FUNCTION_BLOCK "Flag: State Transition"   // FB4, SCL
{ S7_Optimized_Access := 'TRUE' }
VERSION : 0.1
   VAR_IN_OUT
      stns : "Station: All Stations";
   END_VAR
   VAR
      old : Struct
         stn : Array[0.."STATION_COUNT"] of Struct
            orderState : Array[0.."STATION_BUTTON_COUNT"] of Int;
         END_STRUCT;
      END_STRUCT;
   END_VAR
   VAR_TEMP
      pStn : Int;
      pBtn : Int;
      ret : Bool;
   END_VAR
BEGIN
   REGION "FOR EACH STATION"
       FOR #pStn := 0 TO "STATION_COUNT" DO

           REGION "IGNORE WIP LOAD CYCLE"
               IF NOT #stns.stn[#pStn].flags.wipSwapped THEN

                   REGION "FOR EACH BUTTON"
                       FOR #pBtn := 0 TO "STATION_BUTTON_COUNT" DO

                           REGION "RESET RETURN"
                               #ret := FALSE;
                           END_REGION

                           REGION "ON CHANGE IN STATE"
                               IF #stns.stn[#pStn].wipCmpts.orderState[#pBtn] <> #old.stn[#pStn].orderState[#pBtn] THEN

                                   REGION "SET STATE TRANSITION FLAG"
                                       #ret := true;
                                   END_REGION

                               END_IF;
                           END_REGION

                           REGION "SAVE FLAG"
                               #stns.stn[#pStn].flags.stateTransition[#pBtn] := #ret;
                           END_REGION

                       END_FOR;
                   END_REGION

               END_IF;
           END_REGION

           REGION "CHANGE DETECTION"
               #old.stn[#pStn].orderState := #stns.stn[#pStn].wipCmpts.orderState;
           END_REGION

       END_FOR;
   END_REGION
END_FUNCTION_BLOCK

FUNCTION_BLOCK "Flag"   // FB5, SCL
{ S7_Optimized_Access := 'TRUE' }
VERSION : 0.1
   VAR_INPUT
      pnLib : "Recipe: PN Text Library";
   END_VAR
   VAR_IN_OUT
      stns : "Station: All Stations";
      savedStns : "Recipe: HMI Stations Saved Wips";
   END_VAR
   VAR
      "inst New PN Code" : "Flag: New PN Code";
      "inst Flag: State Transition" : "Flag: State Transition";
      "inst Flag: Wip Deselect" : "Flag: Wip Deselect";
      "inst Flag: Wip Swapped" : "Flag: Wip Swapped";
   END_VAR
BEGIN
   REGION "NEW PART NUMBER ASSIGNED"
       #"inst New PN Code"(#stns);
   END_REGION

   REGION "PART NUMBER VALIDATION"
       "Flag: PN Good"(pnLib := #pnLib,
                       stns := #stns);
   END_REGION

   REGION "WIP SWAPPED"
       #"inst Flag: Wip Swapped"(#stns);
   END_REGION

   REGION "STATE TRANSITIONS"
       #"inst Flag: State Transition"(#stns);
   END_REGION

   REGION "WIP DESELECTION"
       #"inst Flag: Wip Deselect"(#savedStns);
   END_REGION
END_FUNCTION_BLOCK

FUNCTION_BLOCK "Flag: Wip Swapped"   // FB10, SCL
{ S7_Optimized_Access := 'TRUE' }
VERSION : 0.1
   VAR_IN_OUT
      stns : "Station: All Stations";
   END_VAR
   VAR
      old : Struct
         wipIndex : Array[0.."STATION_COUNT"] of DInt;
      END_STRUCT;
   END_VAR
   VAR_TEMP
      pStn : Int;
      ret : Bool;
   END_VAR
BEGIN
   REGION "FOR EACH STATION"
       FOR #pStn := 0 TO "STATION_COUNT" DO

           REGION "ON WIP CHANGE"
               IF #stns.stn[#pStn].wipData.index <> #old.wipIndex[#pStn] THEN

                   REGION "SET FLAG"
                       #ret := TRUE;
                   END_REGION

                   REGION "SAVE FLAG"
                       #stns.stn[#pStn].wipCmpts.flags.newPN := #ret;
                   END_REGION

               END_IF;
           END_REGION

           REGION "CHANGE DETECTION"
               #old.wipIndex[#pStn] := #stns.stn[#pStn].wipData.index;
           END_REGION

       END_FOR;
   END_REGION
END_FUNCTION_BLOCK

FUNCTION_BLOCK "Flag: Wip Deselect: Flag Pulse"   // FB17, SCL
{ S7_Optimized_Access := 'TRUE' }
VERSION : 0.1
   VAR_INPUT
      remaining : Real;
      reset : Bool;
   END_VAR
   VAR_IN_OUT
      flag : Bool;
   END_VAR
   VAR RETAIN
      hasBeenFlipped : Bool;
   END_VAR
BEGIN
   #flag := FALSE;

   IF #reset THEN
       #hasBeenFlipped := FALSE;
       RETURN;
   END_IF;

   IF #remaining >= 0.0 THEN
       #hasBeenFlipped := FALSE;
       RETURN;
   END_IF;

   IF NOT #hasBeenFlipped THEN
       IF #remaining < 0.0 THEN
           #hasBeenFlipped := TRUE;
           #flag := TRUE;
       END_IF;
   END_IF;
END_FUNCTION_BLOCK

FUNCTION_BLOCK "Flag: Wip Deselect"   // FB18, SCL
{ S7_Optimized_Access := 'TRUE' }
VERSION : 0.1
   VAR_IN_OUT
      savedStns : "Recipe: HMI Stations Saved Wips";
   END_VAR
   VAR
      "inst Flag Pulses" : Array[0.."STATION_COUNT", 0.."WIP_COUNT"] of "Flag: Wip Deselect: Flag Pulse";
   END_VAR
   VAR_TEMP
      pStn : Int;
      pWip : Int;
   END_VAR
BEGIN
   REGION "FOR EACH STATION"
       FOR #pStn := 0 TO "HMI_STATION_COUNT" DO

           REGION "FOR EACH WIP"
               FOR #pWip := 0 TO "WIP_COUNT" DO

                   REGION "FLAG PULSE"
                       #"inst Flag Pulses"[#pStn, #pWip](remaining := #savedStns.stn[#pStn].wip[#pWip].timers.wdsRemaining,
                                                         flag := #savedStns.stn[#pStn].wip[#pWip].flags.clearWipRequest);
                   END_REGION

               END_FOR;
           END_REGION

       END_FOR;
   END_REGION
END_FUNCTION_BLOCK

FUNCTION "Flag: PN Good" : Void   // FC13, SCL
{ S7_Optimized_Access := 'TRUE' }
VERSION : 0.1
   VAR_INPUT
      pnLib : "Recipe: PN Text Library";
   END_VAR
   VAR_IN_OUT
      stns : "Station: All Stations";
   END_VAR
   VAR_TEMP
      pStn : Int;
      pBtn : Int;
      pnGood : Bool;
   END_VAR
BEGIN
   REGION "FOR EACH STATION"
       FOR #pStn := 0 TO "STATION_COUNT" DO

           REGION "FOR EACH BUTTON"
               FOR #pBtn := 0 TO "STATION_BUTTON_COUNT" DO

                   REGION "ON NEW PN"
                       IF #stns.stn[#pStn].wipCmpts.flags.newPN THEN

                           REGION "VALIDATE PN"
                               #pnGood := "Validate PN"(pnCode := #stns.stn[#pStn].wipCmpts.pnCode[#pBtn],
                                                        pnLib := #pnLib);
                           END_REGION

                           REGION "SAVE TO FLAG"
                               #stns.stn[#pStn].wipCmpts.flags.pnGood[#pBtn] := #pnGood;
                           END_REGION

                       END_IF;
                   END_REGION

               END_FOR;
           END_REGION

       END_FOR;
   END_REGION
END_FUNCTION

// folder: From Excel

FUNCTION_BLOCK "From Excel"   // FB8, SCL
{ S7_Optimized_Access := 'TRUE' }
VERSION : 0.1
   VAR_INPUT
      codeLib : "From Excel: Data";
   END_VAR
   VAR_IN_OUT
      stns : "Station: All Stations";
      svdHMIStnWips : "Recipe: HMI Stations Saved Wips";
   END_VAR
   VAR
      operation_complete : Bool;
      start : Bool;
      states : "Initialize Excel Data: States";
   END_VAR
BEGIN
   REGION "STATE MACHINE"
       "Initialize Excel Data: State Machine"(start := "FirstScan" OR #start,
                                              states := #states,
                                              operation_complete := #operation_complete);
   END_REGION

   REGION "LOAD PART NUMBER CODES TO KP8 STATIONS"
       IF #states.pn_code_to_kp8_station THEN
           "From Excel: PN Code to KP8 Stations"(code_library := #codeLib,
                                                 stations := #stns,
                                                 operation_complete := #operation_complete);
       END_IF;
   END_REGION

   REGION "LOAD PART NUMBER CODES TO SAVED WIPS"
       IF #states.pn_code_to_saved_wips THEN
           "From Excel: PN Code to HMI Station Saved Wips"(code_libarary := #codeLib,
                                                           saved_wip_stations := #svdHMIStnWips,
                                                           operation_complete := #operation_complete);
       END_IF;
   END_REGION

   REGION "LOAD WIP CODES TO SAVED WIPS"
       IF #states.wip_code_to_saved_wips THEN
           "From Excel: Wip Code to HMI Station Saved WIps"(excel_code_library := #codeLib,
                                                            saved_wip_stations := #svdHMIStnWips,
                                                            operation_complete := #operation_complete);
       END_IF;
   END_REGION

   REGION "LOAD ACTIVE WIP TO HMI STATION LIST"
       IF #states.active_wip_to_hmi_station_list THEN
           "From Excel: HMI Stations Load Active WIP"(excel_code_library := #codeLib,
                                                      stations := #stns,
                                                      operation_complete := #operation_complete);
       END_IF;
   END_REGION

   REGION "LOAD ACTIVE WIP TO MASTER STATION LIST"
       IF #states.active_wip_to_master_station_list THEN
           "HMI Station: Load Active WIP into Master Station List"(operation_complete := #operation_complete);
       END_IF;
   END_REGION
END_FUNCTION_BLOCK

FUNCTION "From Excel: PN Code to KP8 Stations" : Void   // FC58, SCL
{ S7_Optimized_Access := 'TRUE' }
VERSION : 0.1
   VAR_INPUT
      code_library : "From Excel: Data";
   END_VAR
   VAR_IN_OUT
      stations : "Station: All Stations";
      operation_complete : Bool;
   END_VAR
   VAR_TEMP
      pointer_source : Int;
      pointer_destination : Int;
   END_VAR
BEGIN
   REGION "KP8 STATIONS
       FOR #pointer_source := 0 TO UDINT_TO_INT("Array.Any.Length"(#code_library.kp8Stns) - 1) DO
           #pointer_destination := #code_library.kp8Stns[#pointer_source].pStn;
           IF #pointer_destination = -1 THEN
               EXIT;
           END_IF;
           #stations.stn[#pointer_destination].wipCmpts.pnCode := #code_library.kp8Stns[#pointer_source].pnCode;
       END_FOR;
       #operation_complete := TRUE;
   END_REGION
END_FUNCTION

FUNCTION "From Excel: PN Code to HMI Station Saved Wips" : Void   // FC61, SCL
{ S7_Optimized_Access := 'TRUE' }
VERSION : 0.1
   VAR_INPUT
      code_libarary : "From Excel: Data";
   END_VAR
   VAR_IN_OUT
      saved_wip_stations : "Recipe: HMI Stations Saved Wips";
      operation_complete : Bool;
   END_VAR
   VAR_TEMP
      pointer_source_station : Int;
      pointer_destination_station : Int;
      pointer_wip : Int;
   END_VAR
BEGIN
   REGION "HMI STATIONS"
       FOR #pointer_source_station := 0 TO UDINT_TO_INT("Array.Any.Length"(#code_libarary.hmiStns) - 1) DO
           #pointer_destination_station := #code_libarary.hmiStns[#pointer_source_station].pStn;
           IF #pointer_destination_station = -1 THEN
               EXIT;
           END_IF;
           FOR #pointer_wip := 0 TO "WIP_COUNT" DO
               #saved_wip_stations.stn[#pointer_source_station].wip[#pointer_wip].pnCode :=
                   #code_libarary.hmiStns[#pointer_source_station].wip[#pointer_wip].pnCode;
           END_FOR;
       END_FOR;
       #operation_complete := TRUE;
   END_REGION
END_FUNCTION

FUNCTION "From Excel: HMI Stations Load Active WIP" : Void   // FC62, SCL
{ S7_Optimized_Access := 'TRUE' }
VERSION : 0.1
   VAR_INPUT
      excel_code_library : "From Excel: Data";
   END_VAR
   VAR_IN_OUT
      stations : "Station: All Stations";
      operation_complete : Bool;
   END_VAR
   VAR_TEMP
      pointer_source : Int;
      pointer_destination : Int;
   END_VAR
BEGIN
   REGION "HMI STATIONS"
       FOR #pointer_source := 0 TO UDINT_TO_INT("Array.Any.Length"(#excel_code_library.hmiStns) - 1) DO
           #pointer_destination := #excel_code_library.hmiStns[#pointer_source].pStn;
           IF #pointer_destination = -1 THEN
               EXIT;
           END_IF;
           #stations.stn[#pointer_destination].wipCmpts.pnCode := #excel_code_library.hmiStns[#pointer_source].wip[0].pnCode;
       END_FOR;
       #operation_complete := TRUE;
   END_REGION
END_FUNCTION

FUNCTION "From Excel: Wip Code to HMI Station Saved WIps" : Void   // FC63, SCL
{ S7_Optimized_Access := 'TRUE' }
VERSION : 0.1
   VAR_INPUT
      excel_code_library : "From Excel: Data";
   END_VAR
   VAR_IN_OUT
      saved_wip_stations : "Recipe: HMI Stations Saved Wips";
      operation_complete : Bool;
   END_VAR
   VAR_TEMP
      "pointer_source _station" : Int;
      pointer_destination_station : Int;
      pointer_wip : Int;
   END_VAR
BEGIN
   REGION "HMI STATIONS"
       FOR #"pointer_source _station" := 0 TO UDINT_TO_INT("Array.Any.Length"(#excel_code_library.hmiStns) - 1) DO
           FOR #pointer_wip := 0 TO "WIP_COUNT" DO
               #saved_wip_stations.stn[#"pointer_source _station"].wip[#pointer_wip].wip.code :=
                   #excel_code_library.hmiStns[#"pointer_source _station"].wip[#pointer_wip].wipCode;
           END_FOR;
       END_FOR;
       #operation_complete := TRUE;
   END_REGION
END_FUNCTION

FUNCTION "Initialize Excel Data: State Machine" : Void   // FC148, SCL
{ S7_Optimized_Access := 'TRUE' }
VERSION : 0.1
   VAR_INPUT
      start : Bool;
   END_VAR
   VAR_IN_OUT
      states : "Initialize Excel Data: States";
      operation_complete : Bool;
   END_VAR
   VAR_TEMP
      clear_states : "Initialize Excel Data: States";
   END_VAR
BEGIN
   REGION "LOAD PART NUMBER CODES TO KP8 STATIONS"
       IF #start AND NOT #operation_complete AND "Initialize Excel Data: All States False"(#states) THEN
           #states := #clear_states;
           #states.pn_code_to_kp8_station := TRUE;
           #operation_complete := FALSE;
       END_IF;
   END_REGION

   REGION "LOAD PART NUMBER CODES TO SAVED WIPS"
       IF #states.pn_code_to_kp8_station AND #operation_complete THEN
           #states := #clear_states;
           #states.pn_code_to_saved_wips := TRUE;
           #operation_complete := FALSE;
       END_IF;
   END_REGION

   REGION "LOAD WIP CODES TO SAVED WIPS"
       IF #states.pn_code_to_saved_wips AND #operation_complete THEN
           #states := #clear_states;
           #states.wip_code_to_saved_wips := TRUE;
           #operation_complete := FALSE;
       END_IF;
   END_REGION

   REGION "LOAD ACTIVE WIP TO HMI STATION LIST"
       IF #states.wip_code_to_saved_wips AND #operation_complete THEN
           #states := #clear_states;
           #states.active_wip_to_hmi_station_list := TRUE;
           #operation_complete := FALSE;
       END_IF;
   END_REGION

   REGION "LOAD ACTIVE WIP TO MASTER STATION LIST"
       IF #states.active_wip_to_hmi_station_list AND #operation_complete THEN
           #states := #clear_states;
           #states.active_wip_to_master_station_list := TRUE;
           #operation_complete := FALSE;
       END_IF;
   END_REGION

   REGION "COMPLETE"
       IF #states.active_wip_to_master_station_list AND #operation_complete THEN
           #states := #clear_states;
           #operation_complete := FALSE;
       END_IF;
   END_REGION
END_FUNCTION

FUNCTION "Initialize Excel Data: All States False" : Bool   // FC149, SCL
{ S7_Optimized_Access := 'TRUE' }
VERSION : 0.1
   VAR_INPUT
      states : "Initialize Excel Data: States";
   END_VAR
   VAR_TEMP
      ret : Bool;
   END_VAR
BEGIN
   IF NOT #states.active_wip_to_hmi_station_list AND
       NOT #states.pn_code_to_kp8_station AND
       NOT #states.active_wip_to_master_station_list AND
       NOT #states.pn_code_to_saved_wips AND
       NOT #states.wip_code_to_saved_wips THEN
       #ret := TRUE;
   END_IF;
   #"Initialize Excel Data: All States False" := #ret;
END_FUNCTION

// folder: Global/Physical

FUNCTION "Physical to Global" : Void   // FC1, LAD
{ S7_Optimized_Access := 'TRUE' }
VERSION : 0.1
   VAR_IN_OUT
      stations : "Station: All Stations";
   END_VAR
   VAR_TEMP
      i : Int;
      kp8In : DWord;
   END_VAR
BEGIN

REGION Network 1 (SCL): MAIN LOOP
   FOR #i := 0 TO "STATION_COUNT" DO

       CASE #i OF
           "VOLVO 16 01":
               #kp8In := "VOLVO 16 01 KP8 In";
           "VOLVO 16 02":
               #kp8In := "VOLVO 16 02 KP8 In";
           "VOLVO 16 03":
               #kp8In := "VOLVO 16 03 KP8 In";
           "VOLVO 16 04":
               #kp8In := "VOLVO 16 04 KP8 In";
           "VOLVO 16 05":
               #kp8In := "VOLVO 16 05 KP8 In";
           "VOLVO 16 06":
               #kp8In := "VOLVO 16 06 KP8 In";
           "VOLVO 16 07":
               #kp8In := "VOLVO 16 07 KP8 In";
           "VOLVO 16 08":
               #kp8In := "VOLVO 16 08 KP8 In";
           "VOLVO 16 09":
               #kp8In := "VOLVO 16 09 KP8 In";
           "VOLVO 16 10":
               #kp8In := "VOLVO 16 10 KP8 In";
           "VOLVO 16 11":
               #kp8In := "VOLVO 16 11 KP8 In";
           "CHM 01":
               #kp8In := "CHM 01 KP8 In";
           "CHM 02":
               #kp8In := "CHM 02 KP8 In";
           "CHM 03":
               #kp8In := "CHM 03 KP8 In";
           "CHM 04":
               #kp8In := "CHM 04 KP8 In";
           "CHM 05":
               #kp8In := "CHM 05 KP8 In";
           "CDO 01":
               #kp8In := "CDO 01 KP8 In";
           "CDO 02":
               #kp8In := "CDO 02 KP8 In";
           "CDO 03":
               #kp8In := "CDO 03 KP8 In";
           "BFL 01":
               #kp8In := "BFL 01 KP8 In";
           "BFL 02":
               #kp8In := "BFL 02 KP8 In";
           "BFL 03":
               #kp8In := "BFL 03 KP8 In";
           "LGS 01":
               #kp8In := "LGS 01 KP8 In";
           "LGS 02":
               #kp8In := "LGS 02 KP8 In";
           "LGS 03":
               #kp8In := "LGS 03 KP8 In";
           "CV 01":
               #kp8In := "CV 01 KP8 In";
           "CV 02":
               #kp8In := "CV 02 KP8 In";
           "CV 03":
               #kp8In := "CV 03 KP8 In";
           "CV 04":
               #kp8In := "CV 04 KP8 In";
           "PC 01":
               #kp8In := "PC 01 KP8 In"; 
           "PC 02":
               #kp8In := "PC 02 KP8 In";
       END_CASE;

       #stations.stn[#i].wipCmpts.ioData.kp8.input := #kp8In.%W1;

   END_FOR;
END_REGION
END_FUNCTION

FUNCTION "Global to Physical" : Void   // FC5, LAD
{ S7_Optimized_Access := 'TRUE' }
VERSION : 0.1
   VAR_IN_OUT
      stations : "Station: All Stations";
   END_VAR
   VAR_TEMP
      i : Int;
      j : Int;
      ET200SP : DWord;
      "KP8 In" : DWord;
      "KP8 Out" : DWord;
      Card : Int;
      stnCount : Int;
   END_VAR
BEGIN

REGION Network 1 (SCL): MAIN LOOP
   FOR #i := 0 TO "STATION_COUNT" DO

       #ET200SP := #stations.stn[#i].wipCmpts.ioData.stkLight;
       #"KP8 Out" := #stations.stn[#i].wipCmpts.ioData.kp8.tempOut;

       CASE #i OF
           "VOLVO 16 01":
               "VOLVO 16 01 IO" := #ET200SP;
               "VOLVO 16 01 KP8 Out" := #"KP8 Out";
           "VOLVO 16 02":
               "VOLVO 16 02 IO" := #ET200SP;
               "VOLVO 16 02 KP8 Out" := #"KP8 Out";
           "VOLVO 16 03":
               "VOLVO 16 03 IO" := #ET200SP;
               "VOLVO 16 03 KP8 Out" := #"KP8 Out";
           "VOLVO 16 04":
               "VOLVO 16 04 IO" := #ET200SP;
               "VOLVO 16 04 KP8 Out" := #"KP8 Out";
           "VOLVO 16 05":
               "VOLVO 16 05 IO" := #ET200SP;
               "VOLVO 16 05 KP8 Out" := #"KP8 Out";
           "VOLVO 16 06":
               "VOLVO 16 06 IO" := #ET200SP;
               "VOLVO 16 06 KP8 Out" := #"KP8 Out";
           "VOLVO 16 07":
               "VOLVO 16 07 IO" := #ET200SP;
               "VOLVO 16 07 KP8 Out" := #"KP8 Out";
           "VOLVO 16 08":
               "VOLVO 16 08 IO" := #ET200SP;
               "VOLVO 16 08 KP8 Out" := #"KP8 Out";
           "VOLVO 16 09":
               "VOLVO 16 09 IO" := #ET200SP;
               "VOLVO 16 09 KP8 Out" := #"KP8 Out";
           "VOLVO 16 10":
               "VOLVO 16 10 IO" := #ET200SP;
               "VOLVO 16 10 KP8 Out" := #"KP8 Out";
           "VOLVO 16 11":
               "VOLVO 16 11 IO" := #ET200SP;
               "VOLVO 16 11 KP8 Out" := #"KP8 Out";
           "CHM 01":
               "CHM 01 IO" := #ET200SP;
               "CHM 01 KP8 Out" := #"KP8 Out";
           "CHM 02":
               "CHM 02 IO" := #ET200SP;
               "CHM 02 KP8 Out" := #"KP8 Out";
           "CHM 03":
               "CHM 03 IO" := #ET200SP;
               "CHM 03 KP8 Out" := #"KP8 Out";
           "CHM 04":
               "CHM 04 IO" := #ET200SP;
               "CHM 04 KP8 Out" := #"KP8 Out";
           "CHM 05":
               "CHM 05 IO" := #ET200SP;
               "CHM 05 KP8 Out" := #"KP8 Out";
           "CDO 01":
               "CDO 01 IO" := #ET200SP;
               "CDO 01 KP8 Out" := #"KP8 Out";
           "CDO 02":
               "CDO 02 IO" := #ET200SP;
               "CDO 02 KP8 Out" := #"KP8 Out";
           "CDO 03":
               "CDO 03 IO" := #ET200SP;
               "CDO 03 KP8 Out" := #"KP8 Out";
           "BFL 01":
               "BFL 01 IO" := #ET200SP;
               "BFL 01 KP8 Out" := #"KP8 Out";
           "BFL 02":
               "BFL 02 IO" := #ET200SP;
               "BFL 02 KP8 Out" := #"KP8 Out";
           "BFL 03":
               "BFL 03 IO" := #ET200SP;
               "BFL 03 KP8 Out" := #"KP8 Out";
           "LGS 01":
               "LGS 01 IO" := #ET200SP;
               "LGS 01 KP8 Out" := #"KP8 Out";
           "LGS 02":
               "LGS 02 IO" := #ET200SP;
               "LGS 02 KP8 Out" := #"KP8 Out";
           "LGS 03":
               "LGS 03 IO" := #ET200SP;
               "LGS 03 KP8 Out" := #"KP8 Out";
           "CV 01":
               "CV 01 IO" := #ET200SP;
               "CV 01 KP8 Out" := #"KP8 Out";
           "CV 02":
               "CV 02 IO" := #ET200SP;
               "CV 02 KP8 Out" := #"KP8 Out";
           "CV 03":
               "CV 03 IO" := #ET200SP;
               "CV 03 KP8 Out" := #"KP8 Out";
           "CV 04":
               "CV 04 IO" := #ET200SP;
               "CV 04 KP8 Out" := #"KP8 Out";
           "PC 01":
               "PC 01 IO" := #ET200SP;
               "PC 01 KP8 Out" := #"KP8 Out";
           "PC 02":
               "PC 02 IO" := #ET200SP;
               "PC 02 KP8 Out" := #"KP8 Out";

       END_CASE;

   END_FOR;
END_REGION
END_FUNCTION

// folder: HMI: Warehouse/001 Part Call

FUNCTION_BLOCK "Part Call"   // FB16, SCL
{ S7_Optimized_Access := 'TRUE' }
VERSION : 0.1
   VAR_INPUT
      tblData : "Part Request Data";
      stns : "Station: All Stations";
      savedWips : "Recipe: HMI Stations Saved Wips";
      pnLib : "Recipe: PN Text Library";
   END_VAR
   VAR_IN_OUT
      tblHMI : "Part Call Screen";
      tableNav : "Nav Bar Data: PLC";
   END_VAR
   VAR RETAIN
      rowIndices : Array[0.."partReqTblHMIRowCnt"] of DInt;
   END_VAR
   VAR
      "inst Table Nav" : "Table Nav";
   END_VAR
   VAR_TEMP
      _tblHMI : "Part Call Screen";
      pRowHMI : DInt;
      pRowData : DInt;
   END_VAR
   // rowIndices[1] := 1;
   // rowIndices[2] := 2;
   // rowIndices[3] := 3;
   // rowIndices[4] := 4;
   // rowIndices[5] := 5;
   // rowIndices[6] := 6;
   // rowIndices[7] := 7;
   // rowIndices[8] := 8;
   // rowIndices[9] := 9;
   // rowIndices[10] := 10;
BEGIN
   REGION "TABLE NAVIGATION"
       #"inst Table Nav"(tblData := #tblData.row,
                         tblDisp := #tblHMI.row,
                         tableNav := #tableNav,
                         rowIndices := #rowIndices);
   END_REGION


   REGION "NAV BUTTON ANIMATIONS"
       "Part Call: Nav Animations"(#tableNav);
   END_REGION

   REGION "DOUBLE BUFFER IN"
       #_tblHMI := #tblHMI;
   END_REGION

   REGION "DRAW HMI TABLE"
       FOR #pRowHMI := 0 TO "partReqTblHMIRowCnt" DO

           REGION "ROW POINTER"
               #pRowData := #rowIndices[#pRowHMI];
           END_REGION

           REGION "DATA"
               "Part Call: Populate HMI Row"(address := #tblData.row[#pRowData],
                                             pnLib := #pnLib,
                                             stns := #stns,
                                             hmiRow := #_tblHMI.row[#pRowHMI]);
           END_REGION

           REGION "ANIMATIONS"
               "Part Call: Row Animations"(address := #tblData.row[#pRowData],
                                           stns := #stns,
                                           savedWips := #savedWips,
                                           rowHMI := #_tblHMI.row[#pRowHMI]);
           END_REGION

       END_FOR;
   END_REGION

   REGION "DOUBLE BUFFER OUT"
       #tblHMI := #_tblHMI;
   END_REGION
END_FUNCTION_BLOCK

FUNCTION "Part Call: Nav Animations" : Void   // FC18, SCL
{ S7_Optimized_Access := 'TRUE' }
VERSION : 0.1
   VAR_IN_OUT
      tableNav : "Nav Bar Data: PLC";
   END_VAR
   VAR_TEMP
      gray : USInt;
      green : USInt;
   END_VAR
BEGIN
   REGION "ANIMATE PART CALL NAV"

       REGION "COPY TO LOCAL"
           #gray := "GRAY_BACKGROUND";
           #green := "GREEN_LIGHT_BACKGROUND";
       END_REGION

       REGION "TOP"
           #tableNav.top.animate := "Bool.Animate"(true_color := #green,
                                                   false_color := #gray,
                                                   evaluation_signal := #tableNav.top.actuate);
       END_REGION

       REGION "PAGE UP"
           #tableNav.pageUp.animate := "Bool.Animate"(true_color := #green,
                                                      false_color := #gray,
                                                      evaluation_signal := #tableNav.pageUp.actuate);
       END_REGION

       REGION "LINE UP"
           #tableNav.lineUp.animate := "Bool.Animate"(true_color := #green,
                                                      false_color := #gray,
                                                      evaluation_signal := #tableNav.lineUp.actuate);
       END_REGION

       REGION "LINE DOWN"
           #tableNav.lineDown.animate := "Bool.Animate"(true_color := #green,
                                                        false_color := #gray,
                                                        evaluation_signal := #tableNav.lineDown.actuate);
       END_REGION

       REGION "PAGE DOWN"
           #tableNav.pageDown.animate := "Bool.Animate"(true_color := #green,
                                                        false_color := #gray,
                                                        evaluation_signal := #tableNav.pageDown.actuate);
       END_REGION

       REGION "BOTTOM"
           #tableNav.bottom.animate := "Bool.Animate"(true_color := #green,
                                                      false_color := #gray,
                                                      evaluation_signal := #tableNav.bottom.actuate);
       END_REGION

   END_REGION
END_FUNCTION

FUNCTION "Part Call: Populate HMI Row" : Void   // FC19, SCL
{ S7_Optimized_Access := 'TRUE' }
VERSION : 0.1
   VAR_INPUT
      address : DInt;
      pnLib : "Recipe: PN Text Library";
      stns : "Station: All Stations";
   END_VAR
   VAR_IN_OUT
      hmiRow : "Table Row";
   END_VAR
   VAR_TEMP
      saveAct : Bool;
      pStn : DInt;
      pWip : DInt;
      pBtn : DInt;
      blankRow : "Table Row";
   END_VAR
BEGIN
   REGION "ROW HAS DATA"
       IF #address <> -1 THEN

           REGION "GET POINTERS"
               #pStn := "Address.Get_Station"(#address);
               #pWip := "Address.Get_Wip"(#address);
               #pBtn := "Address.Get_Button"(#address);
           END_REGION

           REGION "NON WIP SPECIFIC"

           END_REGION

           REGION "GET DATA"
               #hmiRow.address := #address;
               #hmiRow.ordered := "Part Ordered"(#stns.stn[#pStn].wipCmpts.orderState[#pBtn]);
               #hmiRow.tfDropZone.value := "Strip Sign"(USINT_TO_WSTRING(#stns.stn[#pStn].id.dropZone));
               #hmiRow.tfLine.value := #stns.stn[#pStn].id.lineName;
               #hmiRow.tfPartNumber.value := "Part_Number.Code_to_WString"(pnLib := #pnLib, pnCode := #stns.stn[#pStn].wipCmpts.pnCode[#pBtn]);
               #hmiRow.tfTime.value := "Timer.Real_to_WString"(#stns.stn[#pStn].wipCmpts.timers.remaining[#pBtn]);
           END_REGION

       END_IF;
   END_REGION

   REGION "ROW HAS NO DATA"
       IF #address = -1 THEN
           #hmiRow := #blankRow;
       END_IF;
   END_REGION
END_FUNCTION

FUNCTION "Part Call: Row Animations" : Void   // FC20, SCL
{ S7_Optimized_Access := 'TRUE' }
VERSION : 0.1
   VAR_INPUT
      address : DInt;
      stns : "Station: All Stations";
      savedWips : "Recipe: HMI Stations Saved Wips";
   END_VAR
   VAR_IN_OUT
      rowHMI : "Table Row";
   END_VAR
   VAR_TEMP
      cBackground : USInt;
      cForeground : USInt;
      state : Int;
   END_VAR
BEGIN
   REGION "ROW HAS DATA"
       IF #address >= 0 THEN

           REGION "GET STATE"
               #state := "Part Call: Get State"(address := #address,
                                                stns := #stns,
                                                savedWips := #savedWips);
           END_REGION

           REGION "GET COLOR"
               "Part Call: State to Color"(state := #state,
                                           background => #cBackground,
                                           foreground => #cForeground);
           END_REGION

       END_IF;
   END_REGION

   REGION "ROW HAS NO DATA"
       IF #address <= -1 THEN
           #cForeground := "INVISIBLE";
           #cBackground := "INVISIBLE";
       END_IF;
   END_REGION


   REGION "DRAW TO HMI"
       "Part Call: Color Row"(cBackground := #cBackground,
                              cForeground := #cForeground,
                              singleLinePN := TRUE,
                              rowHMI := #rowHMI);
   END_REGION
END_FUNCTION

FUNCTION "Part Call: State to Color" : Void   // FC22, SCL
{ S7_Optimized_Access := 'TRUE' }
VERSION : 0.1
   VAR_INPUT
      state : Int;
   END_VAR
   VAR_OUTPUT
      background : USInt;
      foreground : USInt;
   END_VAR
   VAR_TEMP
      bg : USInt;
      cBlue : USInt;
      cGrayLight : USInt;
      cGrayDark : USInt;
      cGreen : USInt;
      cInvisible : USInt;
      cRedSolid : USInt;
      cRedFlash : USInt;
      cWhite : USInt;
      fg : USInt;
   END_VAR
BEGIN
   #cBlue := "BLUE_LIGHT_BACKGROUND";
   #cGreen := "GREEN_LIGHT_BACKGROUND";
   #cInvisible := "INVISIBLE";
   #cRedSolid := "RED_LIGHT_BACKGROUND";
   #cRedFlash := "RED_LIGHT_FLASHING";
   #cGrayLight := "GRAY_BACKGROUND";
   #cGrayDark := "DISABLED";
   #cWhite := "WHITE_BACKGROUND";

   CASE #state OF
       0, "idle":
           #bg := #cInvisible;
           #fg := #cInvisible;
       "requested", "acknowledged":
           #bg := #cGrayDark;
           #fg := #cGrayLight;
       "requestedCrit", "orderedCrit", "acknowledgedCrit":
           #bg := #cGrayDark;
           #fg := #cRedSolid;
       "requestedExp", "orderedExp", "acknowledgedExp":
           #bg := #cGrayDark;
           #fg := #cRedFlash;
       "ordered":
           #bg := #cGrayDark;
           #fg := #cBlue;
   END_CASE;

   #foreground := #fg;
   #background := #bg;
END_FUNCTION

FUNCTION "Part Call: Color Row" : Void   // FC31, SCL
{ S7_Optimized_Access := 'TRUE' }
VERSION : 0.1
   VAR_INPUT
      cBackground : USInt;
      cForeground : USInt;
      singleLinePN : Bool;
   END_VAR
   VAR_IN_OUT
      rowHMI : "Table Row";
   END_VAR
   VAR_TEMP
      row : "Table Row";
   END_VAR
BEGIN
   REGION "DOUBLE BUFFER IN"
       #row := #rowHMI;
   END_REGION

   REGION "INDEPENDANT ROWS"
       #row.pbSelection.animate := #cForeground;
       #row.rtBackground.animate := #cBackground;
       #row.tfDropZone.animate := #cForeground;
       #row.tfLine.animate := #cForeground;
       #row.tfTime.animate := #cForeground;
   END_REGION


   REGION "DEPENDANT ROWS"

       REGION "SINGLE LINE PART NUMBER"
           IF #singleLinePN THEN
               #row.tfPartNumber.animateDL := "INVISIBLE";
               #row.tfPartNumber.animateSL := #cForeground;
           END_IF;
       END_REGION

       REGION "DOUBLE LINE PN"
           IF NOT #singleLinePN THEN
               #row.tfPartNumber.animateDL := #cForeground;
               #row.tfPartNumber.animateSL := "INVISIBLE";
           END_IF;
       END_REGION

   END_REGION

   REGION "DOUBLE BUFFER OUT"
       #rowHMI := #row;
   END_REGION
END_FUNCTION

FUNCTION "Address in Loaded Wip" : Bool   // FC43, SCL
{ S7_Optimized_Access := 'TRUE' }
VERSION : 0.1
   VAR_INPUT
      pWip : DInt;
      stn : "Station: Single Station";
   END_VAR
   VAR_TEMP
      ret : Bool;
   END_VAR
BEGIN
   IF #pWip = #stn.wipData.index THEN
       #ret := TRUE;
   END_IF;
   #"Address in Loaded Wip" := #ret;
END_FUNCTION

FUNCTION "Part Call: Get State" : Int   // FC57, SCL
{ S7_Optimized_Access := 'TRUE' }
VERSION : 0.1
   VAR_INPUT
      address : DInt;
      stns : "Station: All Stations";
      savedWips : "Recipe: HMI Stations Saved Wips";
   END_VAR
   VAR_TEMP
      addressInWip : Bool;
      pBtn : DInt;
      pStn : DInt;
      pWip : DInt;
      ret : Int;
   END_VAR
BEGIN
   REGION "DECOMPOSE ADDRESS"
       #pBtn := "Address.Get_Button"(#address);
       #pStn := "Address.Get_Station"(#address);
       #pWip := "Address.Get_Wip"(#address);
   END_REGION

   REGION "CHECK ADDRESS AGAINST STATION'S CURRENT WIP"
       #addressInWip := "Address in Loaded Wip"(pWip := #pWip,
                                                stn := #stns.stn[#pStn]);
   END_REGION

   REGION "ADDRESS IN WIP"
       IF #addressInWip THEN
           #ret := #stns.stn[#pStn].wipCmpts.orderState[#pBtn];
       END_IF;
   END_REGION

   REGION "ADDRESS NOT IN WIP"
       IF NOT #addressInWip THEN
           #ret := #savedWips.stn[#pStn].wip[#pWip].orderState[#pBtn];
       END_IF;
   END_REGION

   REGION "RETURN"
       #"Part Call: Get State" := #ret;
   END_REGION
END_FUNCTION

// folder: HMI: Warehouse/002 Settings

FUNCTION_BLOCK "Settings Screen"   // FB19, SCL
{ S7_Optimized_Access := 'TRUE' }
VERSION : 0.1
   VAR_INPUT
      settings_meta : "Setting Meta Data";
      wip_library : "Recipe: Wip Text Library";
   END_VAR
   VAR_IN_OUT
      pn_library : "Recipe: PN Text Library";
      saved_wips : "Recipe: HMI Stations Saved Wips";
      stations : "Station: All Stations";
      settings : "Settings";
   END_VAR
   VAR
      "Assign Button" : "Assign Button";
      "Critical Time IO Field" : "Critical_IO_Field";
      "Dropzone IO Field" : "Dropzone IO Field";
      first_row : DInt;
      "Line IO Field" : "Line IO Field";
      "Part Number IO Field" : "Part Number IO Field";
      process_inputs : "Settings Screen: Processed Inputs";
      "Select Buttons Button" : "Select Buttons";
      "Select Station Button" : "Select Station PB";
      "Select WIP Button" : "Select WIP PB";
      "Table Nav_Instance" : "Table Nav";
      "Total Time IO Field" : "Total_IO_Field";
      "WIP Select Table NavBar" : "NavBar";
      inst_Selected_WIP_Table : "Selected_WIP_Table";
   END_VAR
   VAR_TEMP
      _station_rows_buffer : Array[0..2] of "Settings Station Row Data";
   END_VAR
   VAR CONSTANT
      TABLE_LENGTH : DInt := 49;
      VISIBLE_ROW_COUNT : DInt := 2;
   END_VAR
BEGIN
   REGION "SELECT STATION BUTTON"
       #"Select Station Button"(#settings.selectStation);
   END_REGION

   REGION "SELECT BUTTONS BUTTON"
       #"Select Buttons Button"(settings_meta := #settings_meta,
                                stations := #stations,
                                interface := #settings.selectButton);
   END_REGION

   REGION "SELECT WIP BUTTON"
       #"Select WIP Button"(settings_meta := #settings_meta,
                            stations := #stations,
                            interface := #settings.selectWip);
   END_REGION

   REGION "LINE IO FIELD"
       #"Line IO Field"(settings_meta := #settings_meta,
                        stations := #stations,
                        interface := #settings.line,
                        get_line := #process_inputs.line_name);
   END_REGION

   REGION "DROPZONE IO FIELD"
       #"Dropzone IO Field"(settings_meta := #settings_meta,
                            stations := #stations,
                            interface := #settings.dropzone,
                            get_dropzone := #process_inputs.dropzone);
   END_REGION

   REGION "TOTAL TIME IO FIELD"
       #"Total Time IO Field"(settings_meta := #settings_meta,
                              stations := #stations,
                              interface := #settings.total,
                              state_changes := #process_inputs.total);
   END_REGION

   REGION "CRITICAL TIME IO FIELD"
       #"Critical Time IO Field"(settings_meta := #settings_meta,
                                 stations := #stations,
                                 interface := #settings.critical,
                                 state_changes := #process_inputs.critical);
   END_REGION

   REGION "PART NUMBER ENTRY FIELD"
       #"Part Number IO Field"(settings_meta := #settings_meta,
                               stations := #stations,
                               interface := #settings.partNumber,
                               get_part_number := #process_inputs.part_number_single);

   END_REGION

   REGION "ASSIGN BUTTON"
       #"Assign Button"(critical_time := #settings.critical,
                        drop_zone := #settings.dropzone,
                        line := #settings.line,
                        part_number := #settings.partNumber,
                        settings_meta := #settings_meta,
                        total_time := #settings.total,
                        pn_library := #pn_library,
                        saved_wips := #saved_wips,
                        stations := #stations,
                        interface := #settings.assign,
                        state_changes := #process_inputs.assign);
   END_REGION

   REGION "SELECTED WIP TABLE"
       #_station_rows_buffer := #settings.stationRows;
       #inst_Selected_WIP_Table(saved_wips := #saved_wips,
                                settings_meta := #settings_meta,
                                stations := #stations,
                                wip_library := #wip_library,
                                pn_library := #pn_library,
                                navigation_bar := #settings.stnTableNavBar.plc,
                                stationRows := #_station_rows_buffer);
       #settings.stationRows := #_station_rows_buffer;
   END_REGION

   REGION "WIP SELECT TABLE NAVBAR"
       #"WIP Select Table NavBar"(hide := #settings_meta.selected_stations.count < 4,
                                  TABLE_LENGTH := #TABLE_LENGTH,
                                  VISIBLE_ROW_COUNT := #VISIBLE_ROW_COUNT,
                                  interface := #settings.stnTableNavBar,
                                  first_row := #first_row);
   END_REGION
END_FUNCTION_BLOCK

FUNCTION "Settings Screen: Load Selected: Non-HMI Station" : Void   // FC150, SCL
{ S7_Optimized_Access := 'TRUE' }
VERSION : 0.1
   VAR_INPUT
      stations : "Station: All Stations";
      selected_stations : "Selected Stations";
      wip_library : "Recipe: Wip Text Library";
      part_number_library : "Recipe: PN Text Library";
   END_VAR
   VAR_IN_OUT
      selected_station_table : Array[0..2] of "Settings Station Row Data";
   END_VAR
   VAR_TEMP
      station_index : Int;
      table_row_index : Int;
   END_VAR
BEGIN
   FOR #station_index := 0 TO "STATION_COUNT" DO
       IF #selected_stations.stns[#station_index] THEN
           "Settings Screen: Load Selected WIP"(station := #stations.stn[#station_index],
                                                wip_library := #wip_library,
                                                part_number_library := #part_number_library,
                                                table_row := #selected_station_table[#table_row_index]);
           #table_row_index += 1;
           IF #table_row_index > 2 THEN
               EXIT;
           END_IF;
       END_IF;
   END_FOR;
END_FUNCTION

FUNCTION "Settings Screen: Load Selected WIP" : Void   // FC151, SCL
{ S7_Optimized_Access := 'TRUE' }
VERSION : 0.1
   VAR_INPUT
      station : "Station: Single Station";
      wip_library : "Recipe: Wip Text Library";
      part_number_library : "Recipe: PN Text Library";
   END_VAR
   VAR_IN_OUT
      table_row : "Settings Station Row Data";
   END_VAR
   VAR_TEMP
      _table_row : "Settings Station Row Data";
      button_index : Int;
   END_VAR
BEGIN
   REGION "NOTES"
       (*
       Simple data map from station presented at input to hmi data structure.
       Decision about which data to map is done in parent.
       last edit: 2021-10-06
       *)
   END_REGION

   REGION "BUFFER IN"
       #_table_row := #table_row;
   END_REGION

   REGION "MAP"
       #_table_row.line.data := #station.id.lineName;
       #_table_row.dropzone.data := "Strip Sign"(USINT_TO_WSTRING(#station.id.dropZone));
       #_table_row.wip.data := "WIP.Code_to_WString"(wipTxtLib := #wip_library,
                                                           code := #station.wipData.code);
       FOR #button_index := 0 TO "STATION_BUTTON_COUNT" DO
           "Settings Screen: Load Selected WIP: Load Button"(wip_components:=#station.wipCmpts,
                                                                 wip_library := #wip_library,
                                                                 button_index := #button_index,
                                                                 part_number_liberary := #part_number_library,
                                                                 button_row := #_table_row.btnRows[#button_index]);
       END_FOR;
   END_REGION

   REGION "BUFFER OUT"
       #table_row := #_table_row;
   END_REGION
END_FUNCTION

FUNCTION "Settings Screen: Selected Station Table Row Color" : Void   // FC152, SCL
{ S7_Optimized_Access := 'TRUE' }
VERSION : 0.1
BEGIN
END_FUNCTION

FUNCTION "Settings Screen: Load Selected WIP: Load Button" : Void   // FC155, SCL
{ S7_Optimized_Access := 'TRUE' }
VERSION : 0.1
   VAR_INPUT
      button_index : Int;
      part_number_liberary : "Recipe: PN Text Library";
      wip_components : "Station: Wip: Wip Module";
      wip_library : "Recipe: Wip Text Library";
   END_VAR
   VAR_IN_OUT
      button_row : "Settings Station Row Button Row Data";
   END_VAR
   VAR_TEMP
      _button_row : "Settings Station Row Button Row Data";
      part_number_wstring : WString;
      part_number_code : DInt;
   END_VAR
   VAR CONSTANT
      no_code : WString;
   END_VAR
BEGIN
   REGION "NOTES"
       (*
       Simple data map from station presented at input to hmi data structure.
       Decision about which data to map is done in parent.
       last edit: 2021-10-06
       *)
   END_REGION

   REGION "BUFFER IN"    
       #_button_row := #button_row;
   END_REGION

   REGION "BUTTON LABEL"
       // CURRENTLY A STATIC LABEL
   END_REGION

   REGION "ALOTTED TIME"
       #_button_row.total.data := "Timer.Real_to_WString"(#wip_components.timers.ptAllotted[#button_index]);
   END_REGION

   REGION "CRITICAL TIME"
       #_button_row.critical.data := "Timer.Real_to_WString"(#wip_components.timers.ptCritical[#button_index]);
   END_REGION

   REGION "PART NUMBER"

       REGION "PROCESS PART NUMBER"
           #part_number_code := #wip_components.pnCode[#button_index];
           #part_number_wstring := "Part_Number.Code_to_WString"(pnLib := #part_number_liberary,
                                                         pnCode := #part_number_code);
       END_REGION

       REGION "SINGLE LINE PART NUMBER"
           IF "Part_Number.Is_Single"(#part_number_code) THEN
               #_button_row.singlePN.data := #part_number_wstring;
               #_button_row.doublePN.data := #no_code;
           END_IF;
       END_REGION

       REGION "DOUBLE LINE PART NUMBER"
           IF "Part_Number.Is_Double"(#part_number_code) THEN
               #_button_row.singlePN.data := #no_code;
               #_button_row.doublePN.data := #part_number_wstring;
           END_IF;
       END_REGION

   END_REGION

   REGION "BUFFER OUT"
       #button_row := #_button_row;
   END_REGION
END_FUNCTION

FUNCTION "Settings Screen: Load Selected: HMI Station" : Void   // FC176, SCL
{ S7_Optimized_Access := 'TRUE' }
VERSION : 0.1
   VAR_INPUT
      stations : "Station: All Stations";
      selected_wips : "Selected Wips";
      wip_library : "Recipe: Wip Text Library";
      part_number_library : "Recipe: PN Text Library";
   END_VAR
   VAR_IN_OUT
      selected_station_table : Array[0..2] of "Settings Station Row Data";
   END_VAR
   VAR_TEMP
      station_index : Int;
      table_row_index : Int;
   END_VAR
BEGIN
   FOR #station_index := 0 TO #selected_wips.count DO
       "Settings Screen: Load Selected WIP"(station := #stations.stn[#station_index],
                                            wip_library := #wip_library,
                                            part_number_library := #part_number_library,
                                            table_row := #selected_station_table[#table_row_index]);END_FOR;
END_FUNCTION

// folder: HMI: Warehouse/002 Settings/Assign Button

FUNCTION_BLOCK "Assign Button"   // FB55, SCL
{ S7_Optimized_Access := 'TRUE' }
VERSION : 0.1
   VAR_INPUT
      critical_time : "IO Field Data: Label with Data";
      drop_zone : "IO Field Data: Label with Data";
      line : "IO Field Data: Label with Data";
      part_number : "IO Field Data: Label with Data";
      settings_meta : "Setting Meta Data";
      total_time : "IO Field Data: Label with Data";
   END_VAR
   VAR_IN_OUT
      interface : "Push Button Data";
      pn_library : "Recipe: PN Text Library";
      saved_wips : "Recipe: HMI Stations Saved Wips";
      state_changes : "Push Button Data: State Change Data";
      stations : "Station: All Stations";
   END_VAR
   VAR
      "Push Button: State Changes" : "Push Button: State Changes";
   END_VAR
   VAR_TEMP
      _interface : "Push Button Data";
      _state_changes : "Push Button Data: State Change Data";
   END_VAR
BEGIN
   REGION "BUFFER IN"
       #_interface := #interface;
   END_REGION


   REGION "PROCESS USER INPUT"
       #"Push Button: State Changes"(interface := #_interface,
                                     state_changes := #_state_changes);
   END_REGION


   REGION "ANIMATE"
       "Assign Button: Private: Animate"(settings_meta := #settings_meta,
                                         interface := #_interface);
   END_REGION


   REGION "PERFOM ASSIGNMNET"
       IF #_state_changes.actuate.falling THEN
           "Assign_Button.Perform_Assignment"(critical_time := #critical_time,
                                              drop_zone := #drop_zone,
                                              line := #line,
                                              part_number := #part_number,
                                              settings_meta := #settings_meta,
                                              total_time := #total_time,
                                              pn_library := #pn_library,
                                              stations := #stations,
                                              saved_wips := #saved_wips);
       END_IF;
   END_REGION


   REGION "BUFFER OUT"
       #interface := #_interface;
       #state_changes := #_state_changes;
   END_REGION
END_FUNCTION_BLOCK

FUNCTION "Assign Button: Private: Make Visible / Enable" : Bool   // FC197, SCL
{ S7_Optimized_Access := 'TRUE' }
VERSION : 0.1
   VAR_INPUT
      setting_meta : "Setting Meta Data";
   END_VAR
BEGIN
   #"Assign Button: Private: Make Visible / Enable" :=  #setting_meta.selected_btns.count > 0;
END_FUNCTION

FUNCTION "Assign Button: Private: Animate" : Void   // FC198, SCL
{ S7_Optimized_Access := 'TRUE' }
VERSION : 0.1
   VAR_INPUT
      settings_meta : "Setting Meta Data";
   END_VAR
   VAR_IN_OUT
      interface : "Push Button Data";
   END_VAR
   VAR_TEMP
      selected_station_count : DInt;
   END_VAR
BEGIN
   REGION "COLOR"
   #interface.animate := "WHITE_BACKGROUND";
   END_REGION

   REGION "VISIBILITY
       #interface.visible := "Assign Button: Private: Make Visible / Enable"(setting_meta := #settings_meta);
   END_REGION

   REGION "ENABLE"
       #interface.enable := "Assign Button: Private: Make Visible / Enable"(setting_meta := #settings_meta);
   END_REGION
END_FUNCTION

FUNCTION "Assign_Button.Perform_Assignment" : Void   // FC235, SCL
{ S7_Optimized_Access := 'TRUE' }
VERSION : 0.1
   VAR_INPUT
      critical_time : "IO Field Data: Label with Data";
      drop_zone : "IO Field Data: Label with Data";
      line : "IO Field Data: Label with Data";
      part_number : "IO Field Data: Label with Data";
      settings_meta : "Setting Meta Data";
      total_time : "IO Field Data: Label with Data";
   END_VAR
   VAR_IN_OUT
      pn_library : "Recipe: PN Text Library";
      stations : "Station: All Stations";
      saved_wips : "Recipe: HMI Stations Saved Wips";
   END_VAR
   VAR_TEMP
      _station_indices : Array[0.."STATION_COUNT"] of Int;
   END_VAR
BEGIN
   REGION "DO NOTHING ON NO SELECTED STAION"
       IF #settings_meta.selected_stations.count = 0 THEN
           RETURN;
       END_IF;
   END_REGION


   REGION "HMI STATIONS"
       "Selected_Stations.Indices"(selected_stations:=#settings_meta.selected_stations,
                                   selected_stations_indices:=#_station_indices);
       IF "Is_HMI_Station"(#stations.stn[#_station_indices[0]]) THEN
           "Assign_Button.HMI_Stations"(critical_time := #critical_time,
                                        part_number := #part_number,
                                        settings_meta := #settings_meta,
                                        total_time := #total_time,
                                        pn_library := #pn_library,
                                        saved_wips := #saved_wips);
           RETURN;
       END_IF;
   END_REGION


   REGION "KP8 STATIONS"
       "Assign_Button.KP8_Station"(critical_time := #critical_time,
                                   part_number := #part_number,
                                   settings_meta := #settings_meta,
                                   total_time := #total_time,
                                   all_stations := #stations);
       RETURN;
   END_REGION
END_FUNCTION

// folder: HMI: Warehouse/002 Settings/Assign Button/HMI Station

FUNCTION "Assign_Button.HMI_Stations" : Void   // FC236, SCL
{ S7_Optimized_Access := 'TRUE' }
VERSION : 0.1
   VAR_INPUT
      critical_time : "IO Field Data: Label with Data";
      part_number : "IO Field Data: Label with Data";
      settings_meta : "Setting Meta Data";
      total_time : "IO Field Data: Label with Data";
   END_VAR
   VAR_IN_OUT
      pn_library : "Recipe: PN Text Library";
      saved_wips : "Recipe: HMI Stations Saved Wips";
   END_VAR
   VAR_TEMP
      _i : Int;
      _length : Int;
      _selected_stations : Array[0.."STATION_COUNT"] of Int;
      _p_station : Int;
   END_VAR
BEGIN
   REGION "DO NOTHING IF NO STATIONS SELECTED"
       IF #settings_meta.selected_stations.count = 0 THEN
           RETURN;
       END_IF;
   END_REGION


   REGION "GET INDICES OF SELECTED STATIONS"
       "Selected_Stations.Indices"(selected_stations := #settings_meta.selected_stations,
                                   selected_stations_indices := #_selected_stations);

   END_REGION


   REGION "FOR EACH SELECTED STATION"
       #_length := UDINT_TO_INT("Array.Any.Length"(#saved_wips.stn)) - 1;
       FOR #_i := 0 TO #_length DO

           REGION "ASSIGN TO WIP"
               #_p_station := "WIP.Global_Index_to_HMI_Station_Index"(global_index := #_selected_stations[#_i],
                                                                      saved_WIPs := #saved_wips);
               "Assign_Button.HMI_Stations.WIP"(critical_time := #critical_time,
                                                part_number := #part_number,
                                                selected_wips := #settings_meta.selected_wips,
                                                selected_buttons := #settings_meta.selected_btns,
                                                total_time := #total_time,
                                                pn_library := #pn_library,
                                                stations_wips := #saved_wips.stn[#_p_station]);
           END_REGION

       END_FOR;
   END_REGION
END_FUNCTION

